   "84_Setpoints_LIT304_Refill_High" : Real = PLC "84_Setpoints".LIT304_Refill_High, 1 s
   "84_Setpoints_LIT304_Refill_HighHigh" : Real = PLC "84_Setpoints".LIT304_Refill_HighHigh, 1 s
   "84_Setpoints_PIT358_InitialFill_LowLow" : Real = PLC "84_Setpoints".PIT358_InitialFill_LowLow, 1 s
   "84_Setpoints_PIT358_InitialFill_Low" : Real = PLC "84_Setpoints".PIT358_InitialFill_Low, 1 s
   "84_Setpoints_PIT358_InitialFill_High" : Real = PLC "84_Setpoints".PIT358_InitialFill_High, 1 s
   "84_Setpoints_PIT358_InitialFill_HighHigh" : Real = PLC "84_Setpoints".PIT358_InitialFill_HighHigh, 1 s
   "84_Setpoints_PIT358_Refill_LowLow" : Real = PLC "84_Setpoints".PIT358_Refill_LowLow, 1 s
   "19_AUTO_CMNDS_Data_PIT353_CMND_HighHigh" : Real = PLC "12_AI_Data".PIT112In_SCALED, 1 s
   "80_From_HMI_MAN_DQ_138_5" : Bool = PLC "80_From_HMI".MAN_DQ_138_5, 1 s
   "80_From_HMI_MAN_DQ_138_6" : Bool = PLC "80_From_HMI".MAN_DQ_138_6, 1 s
   "80_From_HMI_MAN_DQ_138_7" : Bool = PLC "80_From_HMI".MAN_DQ_138_7, 1 s
   "86_Times_PRE_GCU_TNK_FILL_DLY" : Time = PLC "86_Times".PRE_GCU_TNK_FILL_DLY, 1 s
   "86_Times_GCU_TNK_FILL_MAX_TIME" : Time = PLC "86_Times".GCU_TNK_FILL_MAX_TIME, 1 s
   "86_Times_E400_STRTD_DLY" : Time = PLC "86_Times".E400_STRTD_DLY, 1 s
   "86_Times_E400_RNG_DLY" : Time = PLC "86_Times".E400_RNG_DLY, 1 s
   "86_Times_CV405_OPND_DLY" : Time = PLC "86_Times".CV405_OPND_DLY, 1 s
   "86_Times_CV406_CLSD_DLY" : Time = PLC "86_Times".CV406_CLSD_DLY, 1 s
   "86_Times_E400_STOP_TIME" : Time = PLC "86_Times".E400_STOP_TIME, 1 s
   "86_Times_P303_STOP_TIME" : Time = PLC "86_Times".P303_STOP_TIME, 1 s
   "86_Times_CV341_OPND_DLY" : Time = PLC "86_Times".CV341_OPND_DLY, 1 s
   "86_Times_GCU_TNK_DRN_MAX_TIME" : Time = PLC "86_Times".GCU_TNK_DRN_MAX_TIME, 1 s
   "86_Times_GCU_FLUSH_TIME" : Time = PLC "86_Times".GCU_FLUSH_TIME, 1 s
   "86_Times_POST_FLUSH_DLY" : Time = PLC "86_Times".POST_FLUSH_DLY, 1 s
   "86_Times_CV341_MAX_TRVL_TIME" : Time = PLC "86_Times".CV341_MAX_TRVL_TIME, 1 s
   "86_Times_VLV_CNFG_DN_DLY" : Time = PLC "86_Times".VLV_CNFG_DN_DLY, 1 s
   "86_Times_CV358_MAX_TRVL_TIME" : Time = PLC "86_Times".CV358_MAX_TRVL_TIME, 1 s
   "86_Times_CV407_MAX_TRVL_TIME" : Time = PLC "100_IGG_AUTO_SEQ_DB".CRNT_STEP, 1 s
   "86_Times_CV409_MAX_TRVL_TIME" : Time = PLC "86_Times".CV409_MAX_TRVL_TIME, 1 s
   "86_Times_CV411_MAX_TRVL_TIME" : Time = PLC "86_Times".CV411_MAX_TRVL_TIME, 1 s
   "86_Times_CV441_MAX_TRVL_TIME" : Time = PLC "86_Times".CV441_MAX_TRVL_TIME, 1 s
   "86_Times_PIT416_TRGT_RMP_TIME" : Real = PLC "86_Times".PIT416_TRGT_RMP_TIME, 1 s
   "86_Times_STEP_MAX_TIME_STP_001" : Time = PLC "86_Times".STEP_MAX_TIME_STP_001, 1 s
   "86_Times_STEP_MAX_TIME_STP_005" : Time = PLC "86_Times".STEP_MAX_TIME_STP_005, 1 s
   "86_Times_STEP_MAX_TIME_STP_010" : Time = PLC "86_Times".STEP_MAX_TIME_STP_010, 1 s
   "86_Times_STEP_MAX_TIME_STP_020" : Time = PLC "86_Times".STEP_MAX_TIME_STP_020, 1 s
   "86_Times_STEP_MAX_TIME_STP_030" : Time = PLC "86_Times".STEP_MAX_TIME_STP_030, 1 s
   "86_Times_STEP_MAX_TIME_STP_040" : Time = PLC "86_Times".STEP_MAX_TIME_STP_040, 1 s
   "86_Times_STEP_MAX_TIME_STP_050" : Time = PLC "86_Times".STEP_MAX_TIME_STP_050, 1 s
   "86_Times_STEP_MAX_TIME_STP_060" : Time = PLC "86_Times".STEP_MAX_TIME_STP_060, 1 s
   "86_Times_CV406_MAX_TRVL_TIME" : Time = PLC "86_Times".CV406_MAX_TRVL_TIME, 1 s
   "86_Times_PRE_CV441_OPN_DLY" : Time = PLC "86_Times".PRE_CV441_OPN_DLY, 1 s
   "86_Times_CV441_CLSD_DLY" : Time = PLC "86_Times".CV441_CLSD_DLY, 1 s
   "86_Times_CV441_OPND_DLY" : Time = PLC "86_Times".CV441_OPND_DLY, 1 s
   "80_From_HMI_MAN_DQ_139_0" : Bool = PLC "80_From_HMI".MAN_DQ_139_0, 1 s
   "80_From_HMI_MAN_DQ_139_1" : Bool = PLC "80_From_HMI".MAN_DQ_139_1, 1 s
   "80_From_HMI_MAN_DQ_139_2" : Bool = PLC "80_From_HMI".MAN_DQ_139_2, 1 s
   "80_From_HMI_MAN_DQ_139_3" : Bool = PLC "80_From_HMI".MAN_DQ_139_3, 1 s
   "80_From_HMI_MAN_DQ_139_4" : Bool = PLC "86_Times".STEP_MAX_TIME_STP_160, 1 s
   "80_From_HMI_MAN_DQ_139_5" : Bool = PLC "80_From_HMI".MAN_DQ_139_5, 1 s
   "80_From_HMI_MAN_DQ_139_6" : Bool = PLC "80_From_HMI".MAN_DQ_139_6, 1 s
   "80_From_HMI_MAN_DQ_139_7" : Bool = PLC "80_From_HMI".MAN_DQ_139_7, 1 s
   "16_AQ_Data_R3_SPR_AQ_802" : Real = PLC "16_AQ_Data".R3_SPR_AQ_802, 1 s
   "16_AQ_Data_R3_SPR_AQ_804" : Real = PLC "16_AQ_Data".R3_SPR_AQ_804, 1 s
   "16_AQ_Data_R3_SPR_AQ_806" : Real = PLC "16_AQ_Data".R3_SPR_AQ_806, 1 s
   "80_From_HMI_MAN_AQ_INC_800" : Bool = PLC "80_From_HMI".MAN_AQ_INC_800, 1 s
   "80_From_HMI_MAN_AQ_DEC_800" : Bool = PLC "80_From_HMI".MAN_AQ_DEC_800, 1 s
   "80_From_HMI_MAN_AQ_INC_802" : Bool = PLC "80_From_HMI".MAN_AQ_INC_802, 1 s
   "80_From_HMI_MAN_AQ_DEC_802" : Bool = PLC "80_From_HMI".MAN_AQ_DEC_802, 1 s
   "80_From_HMI_MAN_AQ_INC_804" : Bool = PLC "80_From_HMI".MAN_AQ_INC_804, 1 s
   "80_From_HMI_MAN_AQ_DEC_804" : Bool = PLC "80_From_HMI".MAN_AQ_DEC_804, 1 s
   "80_From_HMI_MAN_AQ_INC_806" : Bool = PLC "80_From_HMI".MAN_AQ_INC_806, 1 s
   "80_From_HMI_MAN_AQ_DEC_806" : Bool = PLC "80_From_HMI".MAN_AQ_DEC_806, 1 s
   "86_Times_P303_STRTD_DLY" : Time = PLC "86_Times".P303_STRTD_DLY, 1 s
   "86_Times_P303_STPD_DLY" : Time = PLC "86_Times".P303_STPD_DLY, 1 s
   "86_Times_P304_STRTD_DLY" : Time = PLC "86_Times".P304_STRTD_DLY, 1 s
   "86_Times_P304_STPD_DLY" : Time = PLC "86_Times".P304_STPD_DLY, 1 s
   "86_Times_P305_STRTD_DLY" : Time = PLC "86_Times".P305_STRTD_DLY, 1 s
   "86_Times_P305_STPD_DLY" : Time = PLC "86_Times".P305_STPD_DLY, 1 s
   "86_Times_CV341_CLSD_DLY" : Time = PLC "86_Times".CV341_CLSD_DLY, 1 s
   "86_Times_CV358_CLSD_DLY" : Time = PLC "86_Times".CV358_CLSD_DLY, 1 s
   "86_Times_CV401_OPND_DLY" : Time = PLC "86_Times".CV401_OPND_DLY, 1 s
   "86_Times_CV401_CLSD_DLY" : Time = PLC "86_Times".CV401_CLSD_DLY, 1 s
   "84_Setpoints_PIT416_Target" : Real = PLC "84_Setpoints".PIT416_Target, 1 s
   "84_Setpoints_PIT416_Low" : Real = PLC "84_Setpoints".PIT416_Low, 1 s
   "84_Setpoints_PIT416_LowLow" : Real = PLC "84_Setpoints".PIT416_LowLow, 1 s
   "84_Setpoints_TIT406_HighHigh" : Real = PLC "84_Setpoints".TIT406_HighHigh, 1 s
   "20_TANKS_IP_DATA_RIO_02_SECOND_TANK_BWT_PH" : Real = PLC "20_TANKS_IP_DATA".RIO_02.SECOND_TANK.BWT_PH, 1 s
   "20_TANKS_IP_DATA_RIO_02_SECOND_TANK_BWT_TEMP" : Real = PLC "20_TANKS_IP_DATA".RIO_02.SECOND_TANK.BWT_TEMP, 1 s
   "20_TANKS_IP_DATA_RIO_02_SECOND_TANK_BWT_LEVEL" : Real = PLC "20_TANKS_IP_DATA".RIO_02.SECOND_TANK.BWT_LEVEL, 1 s
   "2102_TIME_CALCS_DB_TOT_SEQ_HRS_RMNG" : Int = PLC "2102_TIME_CALCS_DB".TOT_SEQ_HRS_RMNG, 1 s
   "2102_TIME_CALCS_DB_TOT_SEQ_MINS_RMNG" : Int = PLC "2102_TIME_CALCS_DB".TOT_SEQ_MINS_RMNG, 1 s
   "2102_TIME_CALCS_DB_PRE_DWELL_TMR_DN" : Bool = PLC "2102_TIME_CALCS_DB".PRE_DWELL_TMR_DN, 1 s
   "2102_TIME_CALCS_DB_DE_OX_TMR_DN" : Bool = PLC "2102_TIME_CALCS_DB".DE_OX_TMR_DN, 1 s
   "2102_TIME_CALCS_DB_DE_OX_SP_TMR_DN" : Bool = PLC "2102_TIME_CALCS_DB".DE_OX_SP_TMR_DN, 1 s
   "2102_TIME_CALCS_DB_DWELL_TMR_DN" : Bool = PLC "2102_TIME_CALCS_DB".DWELL_TMR_DN, 1 s
   "2102_TIME_CALCS_DB_RE_OX_TMR_DN" : Bool = PLC "2102_TIME_CALCS_DB".RE_OX_TMR_DN, 1 s
   "2102_TIME_CALCS_DB_RE_OX_SP_TMR_DN" : Bool = PLC "2102_TIME_CALCS_DB".RE_OX_SP_TMR_DN, 1 s
   "2102_TIME_CALCS_DB_POST_DWELL_TMR_DN" : Bool = PLC "2102_TIME_CALCS_DB".POST_DWELL_TMR_DN, 1 s
   "2102_TIME_CALCS_DB_PRE_DWELL_MINS_RMNG" : Int = PLC "2102_TIME_CALCS_DB".PRE_DWELL_MINS_RMNG, 1 s
   "20_TANKS_IP_DATA_RIO_02_SECOND_TANK_BWT_DO" : Real = PLC "20_TANKS_IP_DATA".RIO_02.SECOND_TANK.BWT_DO, 1 s
   "2100_AUTO_SEQ_DB_SEQ_RNG" : Bool = PLC "2100_AUTO_SEQ_DB".SEQ_RNG, 1 s
   "2102_TIME_CALCS_DB_DWELL_MINS_RMNG" : Int = PLC "2102_TIME_CALCS_DB".DWELL_MINS_RMNG, 1 s
   "2102_TIME_CALCS_DB_DE_OX_SP_MINS_RMNG" : Int = PLC "2102_TIME_CALCS_DB".DE_OX_SP_MINS_RMNG, 1 s
   "2102_TIME_CALCS_DB_RE_OX_MINS_RMNG" : Int = PLC "2102_TIME_CALCS_DB".RE_OX_MINS_RMNG, 1 s
   "2102_TIME_CALCS_DB_RE_OX_SP_MINS_RMNG" : Int = PLC "2102_TIME_CALCS_DB".RE_OX_SP_MINS_RMNG, 1 s
   "2102_TIME_CALCS_DB_POST_DWELL_MINS_RMNG" : Int = PLC "2102_TIME_CALCS_DB".POST_DWELL_MINS_RMNG, 1 s
   "10_DI_DATA_P_303_ENBLD" : Bool = PLC "10_DI_DATA".P_303_ENBLD, 1 s
   "10_DI_DATA_P_304_ENBLD" : Bool = PLC "10_DI_DATA".P_304_ENBLD, 1 s
   "12_AI_Data_CV_405_SCALED" : Real = PLC "12_AI_Data".CV_405_SCALED, 1 s
   "10_DI_DATA_P_303_OK" : Bool = PLC "10_DI_DATA".P_303_OK, 1 s
   "10_DI_DATA_P_304_OK" : Bool = PLC "10_DI_DATA".P_304_OK, 1 s
   "16_AQ_Data_CV405_CNTRL" : Real = PLC "16_AQ_Data".CV405_CNTRL, 1 s
   "10_DI_DATA_CV358_CLSD" : Bool = PLC "10_DI_DATA".CV358_CLSD, 1 s
   "10_DI_DATA_E_400_RUN" : Bool = PLC "10_DI_DATA".E_400_RUN, 1 s
   "2102_TIME_CALCS_DB_DE_OX_MINS_RMNG" : Int = PLC "2102_TIME_CALCS_DB".DE_OX_MINS_RMNG, 1 s
   "20_TANKS_IP_DATA_RIO_02_FIRST_TANK_BWT_LEVEL" : Real = PLC "20_TANKS_IP_DATA".RIO_02.FIRST_TANK.BWT_LEVEL, 1 s
   "20_TANKS_IP_DATA_RIO_02_FIRST_TANK_BWT_TEMP" : Real = PLC "20_TANKS_IP_DATA".RIO_02.FIRST_TANK.BWT_TEMP, 1 s
   "20_TANKS_IP_DATA_RIO_02_FIRST_TANK_BWT_PH" : Real = PLC "20_TANKS_IP_DATA".RIO_02.FIRST_TANK.BWT_PH, 1 s
   "80_From_HMI_RUN_BTCS" : Bool = PLC "80_From_HMI".RUN_BTCS, 1 s
   "80_From_HMI_RUN_BWTS" : Bool = PLC "80_From_HMI".RUN_BWTS, 1 s
   "2110_BTCS_CNTRL_DB_PRE_DWELL_HRS" : Int = PLC "2110_BTCS_CNTRL_DB".PRE_DWELL_HRS, 1 s
   "2110_BTCS_CNTRL_DB_DE_OX_HRS" : Int = PLC "2110_BTCS_CNTRL_DB".DE_OX_HRS, 1 s
   "2110_BTCS_CNTRL_DB_DE_OX_SP_HRS" : Int = PLC "2110_BTCS_CNTRL_DB".DE_OX_SP_HRS, 1 s
   "2110_BTCS_CNTRL_DB_DWELL_HRS" : Int = PLC "2110_BTCS_CNTRL_DB".DWELL_HRS, 1 s
   "2110_BTCS_CNTRL_DB_RE_OX_HRS" : Int = PLC "2110_BTCS_CNTRL_DB".RE_OX_HRS, 1 s
   "2110_BTCS_CNTRL_DB_RE_OX_SP_HRS" : Int = PLC "2110_BTCS_CNTRL_DB".RE_OX_SP_HRS, 1 s
   "2110_BTCS_CNTRL_DB_POST_DWELL_HRS" : Int = PLC "2110_BTCS_CNTRL_DB".POST_DWELL_HRS, 1 s
   "2110_BTCS_CNTRL_DB_PRE_DWELL_MINS" : Int = PLC "2110_BTCS_CNTRL_DB".PRE_DWELL_MINS, 1 s
   "2110_BTCS_CNTRL_DB_DE_OX_MINS" : Int = PLC "2110_BTCS_CNTRL_DB".DE_OX_MINS, 1 s
   "2110_BTCS_CNTRL_DB_DE_OX_SP_MINS" : Int = PLC "2110_BTCS_CNTRL_DB".DE_OX_SP_MINS, 1 s
   "2110_BTCS_CNTRL_DB_DWELL_MINS" : Int = PLC "2110_BTCS_CNTRL_DB".DWELL_MINS, 1 s
   "2110_BTCS_CNTRL_DB_RE_OX_MINS" : Int = PLC "2110_BTCS_CNTRL_DB".RE_OX_MINS, 1 s
   "2110_BTCS_CNTRL_DB_RE_OX_SP_MINS" : Int = PLC "2110_BTCS_CNTRL_DB".RE_OX_SP_MINS, 1 s
   "2110_BTCS_CNTRL_DB_POST_DWELL_MINS" : Int = PLC "2110_BTCS_CNTRL_DB".POST_DWELL_MINS, 1 s
   "2110_BTCS_CNTRL_DB_TOT_SEQ_HRS" : Int = PLC "2110_BTCS_CNTRL_DB".TOT_SEQ_HRS, 1 s
   "2110_BTCS_CNTRL_DB_TOT_SEQ_MINS" : Int = PLC "2110_BTCS_CNTRL_DB".TOT_SEQ_MINS, 1 s
   "2110_BTCS_CNTRL_DB_RMNG_SEQ_HRS" : Int = PLC "2110_BTCS_CNTRL_DB".RMNG_SEQ_HRS, 1 s
   "2110_BTCS_CNTRL_DB_RMNG_SEQ_MINS" : Int = PLC "2110_BTCS_CNTRL_DB".RMNG_SEQ_MINS, 1 s
   "2110_BTCS_CNTRL_DB_BTCS_STATE" : Int = PLC "2110_BTCS_CNTRL_DB".BTCS_STATE, 1 s
   "2110_BTCS_CNTRL_DB_BTCS_STEP" : Int = PLC "2110_BTCS_CNTRL_DB".BTCS_STEP, 1 s
   "2110_BTCS_CNTRL_DB_START_SEQ" : Bool = PLC "2110_BTCS_CNTRL_DB".START_SEQ, 1 s
   "2110_BTCS_CNTRL_DB_STOP_SEQ" : Bool = PLC "2110_BTCS_CNTRL_DB".STOP_SEQ, 1 s
   "2102_TIME_CALCS_DB_TIMES_VALID" : Bool = PLC "2102_TIME_CALCS_DB".TIMES_VALID, 1 s
   "2110_BTCS_CNTRL_DB_PORT_TANK_STS" : Bool = PLC "2110_BTCS_CNTRL_DB".PORT_TANK_STS, 1 s
   "2110_BTCS_CNTRL_DB_RESET_ALL" : Bool = PLC "2110_BTCS_CNTRL_DB".RESET_ALL, 1 s
   "2110_BTCS_CNTRL_DB_STBD_TANK_STS" : Bool = PLC "2110_BTCS_CNTRL_DB".STBD_TANK_STS, 1 s
   "20_TANKS_IP_DATA_RIO_02_FIRST_TANK_BWT_DO" : Real = PLC "20_TANKS_IP_DATA".RIO_02.FIRST_TANK.BWT_DO, 1 s
   "10_DI_DATA_CV341_CLSD" : Bool = PLC "10_DI_DATA".CV341_CLSD, 1 s
   "86_Times_STEP_MAX_TIME_STP_070" : Time = PLC "86_Times".STEP_MAX_TIME_STP_070, 1 s
   "10_DI_DATA_CV341_OPN" : Bool = PLC "10_DI_DATA".CV341_OPN, 1 s
   "10_DI_DATA_CV411_OPN" : Bool = PLC "10_DI_DATA".CV411_OPN, 1 s
   "84_Setpoints_E400_TT002_HighHigh" : Real = PLC "84_Setpoints".E400_TT002_HighHigh, 1 s
   "84_Setpoints_E400_PT002_HighHigh" : Real = PLC "84_Setpoints".E400_PT002_HighHigh, 1 s
   "19_AUTO_CMNDS_Data_CV405_PID_MDLTG" : Bool = PLC "19_AUTO_CMNDS_Data".CV405_PID_MDLTG, 1 s
   "84_Setpoints_PIT416_HighHigh" : Real = PLC "84_Setpoints".PIT416_HighHigh, 1 s
   "1405_PID_CV405_CtrlParamsBackUp_Gain" : Real = PLC "1405_PID_CV405".CtrlParamsBackUp.Gain, 1 s
   "1405_PID_CV405_CtrlParamsBackUp_Ti" : Real = PLC "1405_PID_CV405".CtrlParamsBackUp.Ti, 1 s
   "10_DI_DATA_R3_SPR_DI_136_0" : Bool = PLC "10_DI_DATA".R3_SPR_DI_136_0, 1 s
   "10_DI_DATA_R3_SPR_DI_136_1" : Bool = PLC "10_DI_DATA".R3_SPR_DI_136_1, 1 s
   "10_DI_DATA_PB_10S1" : Bool = PLC "10_DI_DATA".PB_10S1, 1 s
   "10_DI_DATA_PB_10S2" : Bool = PLC "10_DI_DATA".PB_10S2, 1 s
   "10_DI_DATA_EPB_8S1" : Bool = PLC "10_DI_DATA".EPB_8S1, 1 s
   "10_DI_DATA_E_400_STPD" : Bool = PLC "10_DI_DATA".E_400_STPD, 1 s
   "10_DI_DATA_5T1_PWR_OK" : Bool = PLC "10_DI_DATA".5T1_PWR_OK, 1 s
   "140_PGC_HRS_RUN_DB_SHRS_IP" : Int = PLC "140_PGC_HRS_RUN_DB".SHRS_IP, 1 s
   "10_DI_DATA_6Q6_PWR_OK" : Bool = PLC "10_DI_DATA".6Q6_PWR_OK, 1 s
   "12_AI_Data_SL_400_SCALED" : Real = PLC "12_AI_Data".SL_400_SCALED, 1 s
   "12_AI_Data_R3_SPR_AI_824_SCALED" : Real = PLC "12_AI_Data".R3_SPR_AI_824_SCALED, 1 s
   "12_AI_Data_R3_SPR_AI_826_SCALED" : Real = PLC "12_AI_Data".R3_SPR_AI_826_SCALED, 1 s
   "12_AI_Data_R3_SPR_AI_828_SCALED" : Real = PLC "12_AI_Data".R3_SPR_AI_828_SCALED, 1 s
   "12_AI_Data_R3_SPR_AI_830_SCALED" : Real = PLC "12_AI_Data".R3_SPR_AI_830_SCALED, 1 s
   "19_AUTO_CMNDS_Data_LIT304_CMND_LowLow" : Real = PLC "19_AUTO_CMNDS_Data".LIT304_CMND_LowLow, 1 s
   "19_AUTO_CMNDS_Data_LIT304_CMND_Low" : Real = PLC "19_AUTO_CMNDS_Data".LIT304_CMND_Low, 1 s
   "19_AUTO_CMNDS_Data_LIT304_CMND_Target" : Real = PLC "19_AUTO_CMNDS_Data".LIT304_CMND_Target, 1 s
   "19_AUTO_CMNDS_Data_LIT304_CMND_High" : Real = PLC "19_AUTO_CMNDS_Data".LIT304_CMND_High, 1 s
   "19_AUTO_CMNDS_Data_LIT304_CMND_HighHigh" : Real = PLC "19_AUTO_CMNDS_Data".LIT304_CMND_HighHigh, 1 s
   "84_Setpoints_TIT408_High" : Real = PLC "84_Setpoints".TIT408_High, 1 s
   "84_Setpoints_TIT408_HighHigh" : Real = PLC "84_Setpoints".TIT408_HighHigh, 1 s
   "84_Setpoints_TIT406_High" : Real = PLC "84_Setpoints".TIT406_High, 1 s
   "12_AI_Data_R3_SPR_AI_802_SCALED" : Real = PLC "12_AI_Data".R3_SPR_AI_802_SCALED, 1 s
   "140_PGC_HRS_RUN_DB_SRV_HRS" : Int = PLC "140_PGC_HRS_RUN_DB".SRV_HRS, 1 s
   "140_PGC_HRS_RUN_DB_HRS" : Int = PLC "140_PGC_HRS_RUN_DB".HRS, 1 s
   "140_PGC_HRS_RUN_DB_MINS" : Int = PLC "140_PGC_HRS_RUN_DB".MINS, 1 s
   "10_DI_DATA_CV407_OPN" : Bool = PLC "10_DI_DATA".CV407_OPN, 1 s
   "10_DI_DATA_CV409_CLSD" : Bool = PLC "10_DI_DATA".CV409_CLSD, 1 s
   "10_DI_DATA_CV409_OPN" : Bool = PLC "10_DI_DATA".CV409_OPN, 1 s
   "10_DI_DATA_CV406_OPN" : Bool = PLC "10_DI_DATA".CV406_OPN, 1 s
   "10_DI_DATA_FS_350_FLW_OK" : Bool = PLC "10_DI_DATA".FS_350_FLW_OK, 1 s
   "12_AI_Data_LIT_304_SCALED" : Real = PLC "12_AI_Data".LIT_304_SCALED, 1 s
   "10_DI_DATA_FS_332 FLW_OK" : Bool = PLC "10_DI_DATA"."FS_332 FLW_OK", 1 s
   "10_DI_DATA_CV406_CLSD" : Bool = PLC "10_DI_DATA".CV406_CLSD, 1 s
   "10_DI_DATA_CV407_CLSD" : Bool = PLC "10_DI_DATA".CV407_CLSD, 1 s
   "12_AI_Data_E_400_PT002_SCALED" : Real = PLC "12_AI_Data".E_400_PT002_SCALED, 1 s
   "12_AI_Data_TIT_406_SCALED" : Real = PLC "12_AI_Data".TIT_406_SCALED, 1 s
   "12_AI_Data_PIT_416_SCALED" : Real = PLC "12_AI_Data".PIT_416_SCALED, 1 s
   "12_AI_Data_PIT_353_SCALED" : Real = PLC "12_AI_Data".PIT_353_SCALED, 1 s
   "12_AI_Data_TIT_408_SCALED" : Real = PLC "12_AI_Data".TIT_408_SCALED, 1 s
   "12_AI_Data_PIT_348_SCALED" : Real = PLC "12_AI_Data".PIT_348_SCALED, 1 s
   "12_AI_Data_PIT_358_SCALED" : Real = PLC "12_AI_Data".PIT_358_SCALED, 1 s
   "12_AI_Data_E_400_TE002_SCALED" : Real = PLC "12_AI_Data".E_400_TE002_SCALED, 1 s
   "10_DI_DATA_LS_303_LO" : Bool = PLC "10_DI_DATA".LS_303_LO, 1 s
   "10_DI_DATA_CV441_CLSD" : Bool = PLC "10_DI_DATA".CV441_CLSD, 1 s
   "10_DI_DATA_CV441_OPN" : Bool = PLC "10_DI_DATA".CV441_OPN, 1 s
   "20_TANKS_IP_DATA_RIO_02_FIRST_TANK_DECK_IG_PRESS" : Real = PLC "20_TANKS_IP_DATA".RIO_02.FIRST_TANK.DECK_IG_PRESS, 1 s
   "86_Times_FS332 Delay" : Time = PLC "86_Times"."FS332 Delay", 1 s
   "84_Setpoints_LIT304_InitialFill_High" : Real = PLC "84_Setpoints".LIT304_InitialFill_High, 1 s
   "84_Setpoints_LIT304_InitialFill_Low" : Real = PLC "84_Setpoints".LIT304_InitialFill_Low, 1 s
   "10_DI_DATA_E_400_NOK" : Bool = PLC "10_DI_DATA".E_400_NOK, 1 s
   "10_DI_DATA_E_400_SHTDN" : Bool = PLC "10_DI_DATA".E_400_SHTDN, 1 s
   "140_PGC_HRS_RUN_DB_RST" : Bool = PLC "140_PGC_HRS_RUN_DB".RST, 1 s
   "140_PGC_HRS_RUN_DB_SRVC" : Bool = PLC "140_PGC_HRS_RUN_DB".SRVC, 1 s
   "140_PGC_HRS_RUN_DB_SECS" : Int = PLC "140_PGC_HRS_RUN_DB".SECS, 1 s
   "10_DI_DATA_CV411_CLSD" : Bool = PLC "10_DI_DATA".CV411_CLSD, 1 s
   "86_Times_STEP_MAX_TIME_STP_080" : Time = PLC "86_Times".STEP_MAX_TIME_STP_080, 1 s
   "10_DI_DATA_CV358_OPN" : Bool = PLC "10_DI_DATA".CV358_OPN, 1 s
   "86_Times_STEP_MAX_TIME_STP_100" : Time = PLC "86_Times".STEP_MAX_TIME_STP_100, 1 s
   "14_DQ_DATA_CV_422_3P" : Bool = PLC "14_DQ_DATA".CV_422_3P, 1 s
   "14_DQ_DATA_CV_421_3S" : Bool = PLC "14_DQ_DATA".CV_421_3S, 1 s
   "14_DQ_DATA_R3_SPR_DQ_138_7" : Bool = PLC "14_DQ_DATA".R3_SPR_DQ_138_7, 1 s
   "14_DQ_DATA_CV_422_4P" : Bool = PLC "14_DQ_DATA".CV_422_4P, 1 s
   "14_DQ_DATA_CV_421_4S" : Bool = PLC "14_DQ_DATA".CV_421_4S, 1 s
   "14_DQ_DATA_CV_422_5P" : Bool = PLC "14_DQ_DATA".CV_422_5P, 1 s
   "14_DQ_DATA_CV_421_5S" : Bool = PLC "14_DQ_DATA".CV_421_5S, 1 s
   "14_DQ_DATA_CV_422_6P" : Bool = PLC "14_DQ_DATA".CV_422_6P, 1 s
   "14_DQ_DATA_CV_421_6S" : Bool = PLC "14_DQ_DATA".CV_421_6S, 1 s
   "14_DQ_DATA_CV_422_APT" : Bool = PLC "14_DQ_DATA".CV_422_APT, 1 s
   "14_DQ_DATA_R3_SPR_DQ_139_7" : Bool = PLC "14_DQ_DATA".R3_SPR_DQ_139_7, 1 s
   "100_GCU_AUTO_SEQ_DB_RNG" : Bool = PLC "100_GCU_AUTO_SEQ_DB".RNG, 1 s
   "60_Alarm_Data_GCU_ALARM_WORD_01" : Word = PLC "60_Alarm_Data".GCU_ALARM_WORD_01 AT %DB60.DBW0, 1 s
   "14_DQ_DATA_CV_421_1S" : Bool = PLC "14_DQ_DATA".CV_421_1S, 1 s
   "60_Alarm_Data_GCU_ALARM_WORD_02" : Word = PLC "60_Alarm_Data".GCU_ALARM_WORD_02 AT %DB60.DBW2, 1 s
   "60_Alarm_Data_GCU_ALARM_WORD_04" : Word = PLC "60_Alarm_Data".GCU_ALARM_WORD_04 AT %DB60.DBW6, 1 s
   "60_Alarm_Data_GCU_ALARM_WORD_05" : Word = PLC "60_Alarm_Data".GCU_ALARM_WORD_05 AT %DB60.DBW8, 1 s
   "60_Alarm_Data_GCU_ALARM_WORD_06" : Word = PLC "60_Alarm_Data".GCU_ALARM_WORD_06 AT %DB60.DBW10, 1 s
   "60_Alarm_Data_GCU_ALARM_WORD_07" : Word = PLC "60_Alarm_Data".GCU_ALARM_WORD_07 AT %DB60.DBW12, 1 s
   "60_Alarm_Data_GCU_ALARM_WORD_08" : Word = PLC "60_Alarm_Data".GCU_ALARM_WORD_08 AT %DB60.DBW14, 1 s
   "60_Alarm_Data_GCU_ALARM_WORD_09" : Word = PLC "60_Alarm_Data".GCU_ALARM_WORD_09 AT %DB60.DBW16, 1 s
   "62_Warning_Data_GCU_WARNING_WORD_01" : Word = PLC "62_Warning_Data".GCU_WARNING_WORD_01 AT %DB62.DBW0, 1 s
   "62_Warning_Data_GCU_WARNING_WORD_02" : Word = PLC "62_Warning_Data".GCU_WARNING_WORD_02 AT %DB62.DBW2, 1 s
   "62_Warning_Data_GCU_WARNING_WORD_03" : Word = PLC "62_Warning_Data".GCU_WARNING_WORD_03 AT %DB62.DBW4, 1 s
   "62_Warning_Data_GCU_WARNING_WORD_04" : Word = PLC "62_Warning_Data".GCU_WARNING_WORD_04 AT %DB62.DBW6, 1 s
   "62_Warning_Data_GCU_WARNING_WORD_05" : Word = PLC "62_Warning_Data".GCU_WARNING_WORD_05 AT %DB62.DBW8, 1 s
   "62_Warning_Data_GCU_WARNING_WORD_06" : Word = PLC "62_Warning_Data".GCU_WARNING_WORD_06 AT %DB62.DBW10, 1 s
   "62_Warning_Data_GCU_WARNING_WORD_07" : Word = PLC "62_Warning_Data".GCU_WARNING_WORD_07 AT %DB62.DBW12, 1 s
   "60_Alarm_Data_GCU_ALARM_WORD_03" : Word = PLC "60_Alarm_Data".GCU_ALARM_WORD_03 AT %DB60.DBW4, 1 s
   "62_Warning_Data_GCU_WARNING_WORD_08" : Word = PLC "62_Warning_Data".GCU_WARNING_WORD_08 AT %DB62.DBW14, 1 s
   "14_DQ_DATA_CV_422_1P" : Bool = PLC "14_DQ_DATA".CV_422_1P, 1 s
   "14_DQ_DATA_E_400_STP" : Bool = PLC "14_DQ_DATA".E_400_STP, 1 s
   "150_GCU_LCL_CNTRL_DB_SYS_OK_FOR_LCL" : Bool = PLC "150_GCU_LCL_CNTRL_DB".SYS_OK_FOR_LCL, 1 s
   "150_GCU_LCL_CNTRL_DB_RUN_WITH_AIR" : Bool = PLC "150_GCU_LCL_CNTRL_DB".RUN_WITH_AIR, 1 s
   "150_GCU_LCL_CNTRL_DB_RUN_WITH_IG" : Bool = PLC "150_GCU_LCL_CNTRL_DB".RUN_WITH_IG, 1 s
   "80_From_HMI_Request_Auto" : Bool = PLC "80_From_HMI".Request_Auto, 1 s
   "80_From_HMI_Request_Manual" : Bool = PLC "80_From_HMI".Request_Manual, 1 s
   "80_From_HMI_RST_AUT_SEQ" : Bool = PLC "80_From_HMI".RST_AUT_SEQ, 1 s
   "141_P303_HRS_RUN_DB_HRS" : Int = PLC "141_P303_HRS_RUN_DB".HRS, 1 s
   "141_P303_HRS_RUN_DB_MINS" : Int = PLC "141_P303_HRS_RUN_DB".MINS, 1 s
   "141_P303_HRS_RUN_DB_SECS" : Int = PLC "141_P303_HRS_RUN_DB".SECS, 1 s
   "141_P303_HRS_RUN_DB_RST" : Bool = PLC "141_P303_HRS_RUN_DB".RST, 1 s
   "141_P303_HRS_RUN_DB_SRV_HRS" : Int = PLC "141_P303_HRS_RUN_DB".SRV_HRS, 1 s
   "141_P303_HRS_RUN_DB_SHRS_IP" : Int = PLC "141_P303_HRS_RUN_DB".SHRS_IP, 1 s
   "141_P303_HRS_RUN_DB_SRVC" : Bool = PLC "141_P303_HRS_RUN_DB".SRVC, 1 s
   "14_DQ_DATA_CV_422_FPT" : Bool = PLC "14_DQ_DATA".CV_422_FPT, 1 s
   "14_DQ_DATA_P_303" : Bool = PLC "14_DQ_DATA".P_303, 1 s
   "142_P304_HRS_RUN_DB_MINS" : Int = PLC "142_P304_HRS_RUN_DB".MINS, 1 s
   "142_P304_HRS_RUN_DB_SECS" : Int = PLC "142_P304_HRS_RUN_DB".SECS, 1 s
   "142_P304_HRS_RUN_DB_RST" : Bool = PLC "142_P304_HRS_RUN_DB".RST, 1 s
   "142_P304_HRS_RUN_DB_SRV_HRS" : Int = PLC "142_P304_HRS_RUN_DB".SRV_HRS, 1 s
   "142_P304_HRS_RUN_DB_SHRS_IP" : Int = PLC "142_P304_HRS_RUN_DB".SHRS_IP, 1 s
   "142_P304_HRS_RUN_DB_SRVC" : Bool = PLC "142_P304_HRS_RUN_DB".SRVC, 1 s
   "14_DQ_DATA_P_304" : Bool = PLC "14_DQ_DATA".P_304, 1 s
   "100_GCU_AUTO_SEQ_DB_CRNT_STEP" : Int = PLC "100_GCU_AUTO_SEQ_DB".CRNT_STEP, 1 s
   "14_DQ_DATA_13P1" : Bool = PLC "14_DQ_DATA".13P1, 1 s
   "14_DQ_DATA_13P2" : Bool = PLC "14_DQ_DATA".13P2, 1 s
   "14_DQ_DATA_13P3" : Bool = PLC "14_DQ_DATA".13P3, 1 s
   "14_DQ_DATA_13P4" : Bool = PLC "14_DQ_DATA".13P4, 1 s
   "14_DQ_DATA_13P5" : Bool = PLC "14_DQ_DATA".13P5, 1 s
   "142_P304_HRS_RUN_DB_HRS" : Int = PLC "142_P304_HRS_RUN_DB".HRS, 1 s
   "62_Warning_Data_GCU_WARNING_WORD_09" : Word = PLC "62_Warning_Data".GCU_WARNING_WORD_09 AT %DB62.DBW16, 1 s
   "2060_Alarm_Data_BTCS_ALARM_WORD_01" : Word = PLC "2060_Alarm_Data".BTCS_ALARM_WORD_01 AT %DB2060.DBW0, 1 s
   "2060_Alarm_Data_BTCS_ALARM_WORD_02" : Word = PLC "2060_Alarm_Data".BTCS_ALARM_WORD_02 AT %DB2060.DBW2, 1 s
   "504_Tank Grouping_DB2020_TANK ACTIV 12" : Bool = PLC "504_Tank Grouping_DB2020"."TANK ACTIV 12" AT %DB1.DBW0, 1 s
   "504_Tank Grouping_DB2020_TANK ACTIV 14" : Bool = PLC "504_Tank Grouping_DB2020"."TANK ACTIV 14" AT %DB1.DBW0, 1 s
   "504_Tank Grouping_DB2020_TANK ACTIV 16" : Bool = PLC "504_Tank Grouping_DB2020"."TANK ACTIV 16" AT %DB1.DBW0, 1 s
   "504_Tank Grouping_DB2020_TANK ACTIV 18" : Bool = PLC "504_Tank Grouping_DB2020"."TANK ACTIV 18" AT %DB1.DBW0, 1 s
   "504_Tank Grouping_DB2020_TANK ACTIV 20" : Bool = PLC "504_Tank Grouping_DB2020"."TANK ACTIV 20" AT %DB1.DBW0, 1 s
   "504_Tank Grouping_DB2020_TANK ACTIV 3" : Bool = PLC "504_Tank Grouping_DB2020"."TANK ACTIV 3" AT %DB1.DBW0, 1 s
   "504_Tank Grouping_DB2020_TANK ACTIV 5" : Bool = PLC "504_Tank Grouping_DB2020"."TANK ACTIV 5" AT %DB1.DBW0, 1 s
   "504_Tank Grouping_DB2020_TANK ACTIV 7" : Bool = PLC "504_Tank Grouping_DB2020"."TANK ACTIV 7" AT %DB1.DBW0, 1 s
   "504_Tank Grouping_DB2020_TANK ACTIV 9" : Bool = PLC "504_Tank Grouping_DB2020"."TANK ACTIV 9" AT %DB1.DBW0, 1 s
   "504_Tank Grouping_DB2020_TANK ACTIV 11" : Bool = PLC "504_Tank Grouping_DB2020"."TANK ACTIV 11" AT %DB1.DBW0, 1 s
   "504_Tank Grouping_DB2020_TANK ACTIV 13" : Bool = PLC "504_Tank Grouping_DB2020"."TANK ACTIV 13" AT %DB1.DBW0, 1 s
   "504_Tank Grouping_DB2020_TANK ACTIV 1" : Bool = PLC "504_Tank Grouping_DB2020"."TANK ACTIV 1" AT %DB1.DBW0, 1 s
   "504_Tank Grouping_DB2020_TANK ACTIV 17" : Bool = PLC "504_Tank Grouping_DB2020"."TANK ACTIV 17" AT %DB1.DBW0, 1 s
   "504_Tank Grouping_DB2020_TANK ACTIV 10" : Bool = PLC "504_Tank Grouping_DB2020"."TANK ACTIV 10" AT %DB1.DBW0, 1 s
   "504_Tank Grouping_DB2020_TANK ACTIV 19" : Bool = PLC "504_Tank Grouping_DB2020"."TANK ACTIV 19" AT %DB1.DBW0, 1 s
   "2110_BTCS_CNTRL_DB_PORT_TANK_STS(1)" : Bool = PLC "2110_BTCS_CNTRL_DB".PORT_TANK_STS AT %DB1.DBX0.0, 1 s
   "2110_BTCS_CNTRL_DB_STBD_TANK_STS(1)" : Bool = PLC "2110_BTCS_CNTRL_DB".STBD_TANK_STS, 1 s
   "2102_TIME_CALCS_DB_PRE-DWEL_Warning 1" : Bool = PLC "2102_TIME_CALCS_DB"."PRE-DWEL_Warning 1", 500 ms
      on ChangeValue: "TimeRemainingToTreatment"()
   "2102_TIME_CALCS_DB_PRE-DWEL_Warning Min 1" : Int = PLC "2102_TIME_CALCS_DB"."PRE-DWEL_Warning Min 1", 1 s
   "2102_TIME_CALCS_DB_PRE-DWEL_Warning Min 2" : Int = PLC "2102_TIME_CALCS_DB"."PRE-DWEL_Warning Min 2", 1 s
   "2102_TIME_CALCS_DB_PRE-DWEL_Warning Min 3" : Int = PLC "2102_TIME_CALCS_DB"."PRE-DWEL_Warning Min 3", 1 s
   "2102_TIME_CALCS_DB_PRE-DWEL_Warning Reset 1" : Bool = PLC "2102_TIME_CALCS_DB"."PRE-DWEL_Warning Reset 1", 1 s
   "2102_TIME_CALCS_DB_PRE-DWEL_Warning 2" : Bool = PLC "2102_TIME_CALCS_DB"."PRE-DWEL_Warning 2", 500 ms
      on ChangeValue: "TreatmentRequired"()
   "2102_TIME_CALCS_DB_PRE-DWEL_Warning 3" : Bool = PLC "2102_TIME_CALCS_DB"."PRE-DWEL_Warning 3", 1 s
   "2102_TIME_CALCS_DB_PRE-DWEL_Warning Reset 2" : Bool = PLC "2102_TIME_CALCS_DB"."PRE-DWEL_Warning Reset 2", 1 s
   "2102_TIME_CALCS_DB_PRE-DWEL_Warning Reset 3" : Bool = PLC "2102_TIME_CALCS_DB"."PRE-DWEL_Warning Reset 3", 1 s
   "2102_TIME_CALCS_DB_60X boost" : Bool = PLC "2102_TIME_CALCS_DB"."60X boost", 1 s
   "86_Times_STEP_MAX_TIME_STP_090" : Time = PLC "86_Times".STEP_MAX_TIME_STP_090, 1 s
   "504_Tank Grouping_DB2020_TANK ACTIV 21" : Bool = PLC "504_Tank Grouping_DB2020"."TANK ACTIV 21" AT %DB1.DBW0, 1 s
   "504_Tank Grouping_DB2020_TANK ACTIV 8" : Bool = PLC "504_Tank Grouping_DB2020"."TANK ACTIV 8" AT %DB1.DBW0, 1 s
   "504_Tank Grouping_DB2020_TANK ACTIV 6" : Bool = PLC "504_Tank Grouping_DB2020"."TANK ACTIV 6" AT %DB1.DBW0, 1 s
   "504_Tank Grouping_DB2020_TANK ACTIV 4" : Bool = PLC "504_Tank Grouping_DB2020"."TANK ACTIV 4" AT %DB1.DBW0, 1 s
   "2060_Alarm_Data_BTCS_ALARM_WORD_03" : Word = PLC "2060_Alarm_Data".BTCS_ALARM_WORD_03 AT %DB2060.DBW4, 1 s
   "2060_Alarm_Data_BTCS_ALARM_WORD_04" : Word = PLC "2060_Alarm_Data".BTCS_ALARM_WORD_04 AT %DB2060.DBW6, 1 s
   "2060_Alarm_Data_BTCS_ALARM_WORD_05" : Word = PLC "2060_Alarm_Data".BTCS_ALARM_WORD_05 AT %DB2060.DBW8, 1 s
   "2060_Alarm_Data_BTCS_ALARM_WORD_06" : Word = PLC "2060_Alarm_Data".BTCS_ALARM_WORD_06 AT %DB2060.DBW10, 1 s
   "2060_Alarm_Data_BTCS_ALARM_WORD_07" : Word = PLC "2060_Alarm_Data".BTCS_ALARM_WORD_07 AT %DB2060.DBW12, 1 s
   "2060_Alarm_Data_BTCS_ALARM_WORD_08" : Word = PLC "2060_Alarm_Data".BTCS_ALARM_WORD_08 AT %DB2060.DBW14, 1 s
   "80_From_HMI_SAL_VALUE" : Real = PLC "80_From_HMI".SAL_VALUE, 1 s
   "80_From_HMI_SAL_CNFRM" : Bool = PLC "80_From_HMI".SAL_CNFRM, 1 s
   "150_GCU_LCL_CNTRL_DB_OPN_ACTV_GTT_VLVS" : Bool = PLC "150_GCU_LCL_CNTRL_DB".OPN_ACTV_GTT_VLVS, 1 s
   "2068_Sys_Status_Data_SAL_CNF_CHK" : Bool = PLC "2068_Sys_Status_Data".SAL_CNF_CHK, 100 ms
      on ChangeValue: "Salinity_FreshWaterAlert"()
   "80_From_HMI_LOW_SAL_ACPT" : Bool = PLC "80_From_HMI".LOW_SAL_ACPT, 1 s
   "80_From_HMI_LOW_SAL_RJCT" : Bool = PLC "80_From_HMI".LOW_SAL_RJCT, 1 s
   "86_Times_PIT353 Delay" : Time = PLC "86_Times"."PIT353 Delay", 1 s
   "86_Times_PIT416 Delay" : Time = PLC "86_Times"."PIT416 Delay", 1 s
   "19_AUTO_CMNDS_Data_PIT416_CMND_Target" : Real = PLC "19_AUTO_CMNDS_Data".PIT416_CMND_Target, 1 s
   "2102_TIME_CALCS_DB_Voyage_TIME_days" : Int = PLC "2102_TIME_CALCS_DB".Voyage_TIME_days, 1 s
   "2102_TIME_CALCS_DB_Voyage_TIME_invalid" : Bool = PLC "2102_TIME_CALCS_DB".Voyage_TIME_invalid AT %DB1.DBW0, 1 s
      on ChangeValue: "VoyageTimeInsufficient"()
   "2102_TIME_CALCS_DB_TOT_SEQ_DAYS" : Real = PLC "2102_TIME_CALCS_DB".TOT_SEQ_DAYS, 1 s
   "2102_TIME_CALCS_DB_POST_DWELL_TMR_DN(1)" : Bool = PLC "2102_TIME_CALCS_DB".POST_DWELL_TMR_DN AT %DB1.DBD0, 1 s
   "2102_TIME_CALCS_DB_PRE-DWEL HOURS REMNG" : Int = PLC "2102_TIME_CALCS_DB"."PRE-DWEL HOURS REMNG" AT %DB1.DBW0, 1 s
   "504_Tank Grouping_DB2020_TANK ACTIV 2" : Bool = PLC "504_Tank Grouping_DB2020"."TANK ACTIV 2" AT %DB1.DBW0, 1 s
   "150_GCU_LCL_CNTRL_DB_STOP" : Bool = PLC "150_GCU_LCL_CNTRL_DB".STOP, 1 s
   "150_GCU_LCL_CNTRL_DB_STRT_IG" : Bool = PLC "150_GCU_LCL_CNTRL_DB".STRT_IG, 1 s
   "2068_Sys_Status_Data_SAL_VALID" : Bool = PLC "2068_Sys_Status_Data".SAL_VALID, 1 s
   "504_Tank Grouping_DB2020_Sequence Time m Offset_Real" : Real = PLC "504_Tank Grouping_DB2020"."Sequence Time m Offset_real", 1 s
   "86_Times_STEP_MAX_TIME_STP_410" : Time = PLC "86_Times".STEP_MAX_TIME_STP_410, 1 s
   "86_Times_STEP_MAX_TIME_STP_420" : Time = PLC "86_Times".STEP_MAX_TIME_STP_420, 1 s
   "86_Times_STEP_MAX_TIME_STP_430" : Time = PLC "86_Times".STEP_MAX_TIME_STP_430, 1 s
   "86_Times_STEP_MAX_TIME_STP_440" : Time = PLC "86_Times".STEP_MAX_TIME_STP_440, 1 s
   "86_Times_STEP_MAX_TIME_STP_450" : Time = PLC "86_Times".STEP_MAX_TIME_STP_450, 1 s
   "86_Times_STEP_MAX_TIME_STP_460" : Time = PLC "86_Times".STEP_MAX_TIME_STP_460, 1 s
   "86_Times_STEP_MAX_TIME_STP_470" : Time = PLC "86_Times".STEP_MAX_TIME_STP_470, 1 s
   "86_Times_STEP_MAX_TIME_STP_480" : Time = PLC "86_Times".STEP_MAX_TIME_STP_480, 1 s
   "86_Times_STEP_MAX_TIME_STP_490" : Time = PLC "86_Times".STEP_MAX_TIME_STP_490, 1 s
   "86_Times_STEP_MAX_TIME_STP_500" : Time = PLC "86_Times".STEP_MAX_TIME_STP_500, 1 s
   "86_Times_STEP_MAX_TIME_STP_510" : Time = PLC "86_Times".STEP_MAX_TIME_STP_510, 1 s
   "86_Times_STEP_MAX_TIME_STP_520" : Time = PLC "86_Times".STEP_MAX_TIME_STP_520, 1 s
   "86_Times_STEP_MAX_TIME_STP_530" : Time = PLC "86_Times".STEP_MAX_TIME_STP_530, 1 s
   "86_Times_STEP_MAX_TIME_STP_540" : Time = PLC "86_Times".STEP_MAX_TIME_STP_540, 1 s
   "86_Times_STEP_MAX_TIME_STP_550" : Time = PLC "86_Times".STEP_MAX_TIME_STP_550, 1 s
   "86_Times_STEP_MAX_TIME_STP_560" : Time = PLC "86_Times".STEP_MAX_TIME_STP_560, 1 s
   "86_Times_STEP_MAX_TIME_STP_570" : Time = PLC "86_Times".STEP_MAX_TIME_STP_570, 1 s
   "86_Times_STEP_MAX_TIME_STP_580" : Time = PLC "86_Times".STEP_MAX_TIME_STP_580, 1 s
   "86_Times_STEP_MAX_TIME_STP_590" : Time = PLC "86_Times".STEP_MAX_TIME_STP_590, 1 s
   "86_Times_STEP_MAX_TIME_STP_600" : Time = PLC "86_Times".STEP_MAX_TIME_STP_600, 1 s
   "86_Times_STEP_MAX_TIME_STP_610" : Time = PLC "86_Times".STEP_MAX_TIME_STP_610, 1 s
   "86_Times_STEP_MAX_TIME_STP_620" : Time = PLC "86_Times".STEP_MAX_TIME_STP_620, 1 s
   "86_Times_STEP_MAX_TIME_STP_630" : Time = PLC "86_Times".STEP_MAX_TIME_STP_630, 1 s
   "20_TANKS_IP_DATA_RIO_02_FIRST_TANK_TANK_VENT_A_OPEN" : Bool = PLC "20_TANKS_IP_DATA".RIO_02.FIRST_TANK.TANK_VENT_A_OPEN AT %DB1.DBW0, 1 s
   "40_TANKS_OP_DATA_RIO_02_VENT_A_2P" : Bool = PLC "40_TANKS_OP_DATA".RIO_02_VENT_A_2P AT %DB1.DBW0, 1 s
   "86_Times_STEP_MAX_TIME_STP_400" : Time = PLC "86_Times".STEP_MAX_TIME_STP_400, 1 s
   "86_Times_STEP_MAX_TIME_STP_390" : Time = PLC "86_Times".STEP_MAX_TIME_STP_390, 1 s
   "86_Times_STEP_MAX_TIME_STP_380" : Time = PLC "86_Times".STEP_MAX_TIME_STP_380, 1 s
   "86_Times_STEP_MAX_TIME_STP_370" : Time = PLC "86_Times".STEP_MAX_TIME_STP_370, 1 s
   "86_Times_STEP_MAX_TIME_STP_110" : Time = PLC "86_Times".STEP_MAX_TIME_STP_110, 1 s
   "150_GCU_LCL_CNTRL_DB_STRT_AIR" : Bool = PLC "150_GCU_LCL_CNTRL_DB".STRT_AIR, 1 s
   "86_Times_STEP_MAX_TIME_STP_120" : Time = PLC "86_Times".STEP_MAX_TIME_STP_120, 1 s
   "86_Times_STEP_MAX_TIME_STP_130" : Time = PLC "86_Times".STEP_MAX_TIME_STP_001, 1 s
   "86_Times_STEP_MAX_TIME_STP_140" : Time = PLC "86_Times".STEP_MAX_TIME_STP_140, 1 s
   "86_Times_STEP_MAX_TIME_STP_150" : Time = PLC "86_Times".STEP_MAX_TIME_STP_150, 1 s
   "86_Times_STEP_MAX_TIME_STP_160" : Time = PLC "86_Times".STEP_MAX_TIME_STP_160, 1 s
   "86_Times_STEP_MAX_TIME_STP_170" : Time = PLC "86_Times".STEP_MAX_TIME_STP_170, 1 s
   "86_Times_STEP_MAX_TIME_STP_180" : Time = PLC "86_Times".STEP_MAX_TIME_STP_180, 1 s
   "86_Times_STEP_MAX_TIME_STP_190" : Time = PLC "86_Times".STEP_MAX_TIME_STP_190, 1 s
   "86_Times_STEP_MAX_TIME_STP_200" : Time = PLC "86_Times".STEP_MAX_TIME_STP_200, 1 s
   "86_Times_STEP_MAX_TIME_STP_210" : Time = PLC "86_Times".STEP_MAX_TIME_STP_210, 1 s
   "20_TANKS_IP_DATA_RIO_02_FIRST_TANK_GTT_ISOL_VALVE_OPEN" : Bool = PLC "20_TANKS_IP_DATA".RIO_02.FIRST_TANK.GTT_ISOL_VALVE_OPEN AT %DB1.DBW0, 1 s
   "86_Times_STEP_MAX_TIME_STP_220" : Time = PLC "86_Times".STEP_MAX_TIME_STP_220, 1 s
   "86_Times_STEP_MAX_TIME_STP_240" : Time = PLC "86_Times".STEP_MAX_TIME_STP_240, 1 s
   "86_Times_STEP_MAX_TIME_STP_250" : Time = PLC "86_Times".STEP_MAX_TIME_STP_250, 1 s
   "86_Times_STEP_MAX_TIME_STP_260" : Time = PLC "86_Times".STEP_MAX_TIME_STP_260, 1 s
   "86_Times_STEP_MAX_TIME_STP_270" : Time = PLC "86_Times".STEP_MAX_TIME_STP_270, 1 s
   "86_Times_STEP_MAX_TIME_STP_280" : Time = PLC "86_Times".STEP_MAX_TIME_STP_280, 1 s
   "86_Times_STEP_MAX_TIME_STP_290" : Time = PLC "86_Times".STEP_MAX_TIME_STP_290, 1 s
   "86_Times_STEP_MAX_TIME_STP_300" : Time = PLC "86_Times".STEP_MAX_TIME_STP_300, 1 s
   "86_Times_STEP_MAX_TIME_STP_310" : Time = PLC "86_Times".STEP_MAX_TIME_STP_310, 1 s
   "86_Times_STEP_MAX_TIME_STP_320" : Time = PLC "86_Times".STEP_MAX_TIME_STP_320, 1 s
   "86_Times_STEP_MAX_TIME_STP_330" : Time = PLC "86_Times".STEP_MAX_TIME_STP_330, 1 s
   "86_Times_STEP_MAX_TIME_STP_340" : Time = PLC "86_Times".STEP_MAX_TIME_STP_340, 1 s